// Mitsubishi GX Works2 project: 40国轩高温2次注液尝试优化   PLC: Q06UDEH (continued)
CASE iStep OF
	0:(*//初始化*)
	ConveyorMotor.xMotorCW:=0;
	ConveyorMotor.xMotorCCW:=0;
	ConveyorMotor.iProductCategoryOut:=0;
(*	//判断物料有无传感器*)	
		IF m_xPresentDelay THEN			
			ConveyorMotor.xEmpty:=0;
			IF g_xAuto AND NOT ConveyorMotor.xError THEN(*//自动情况下进行跳转*)(*无超限报警*)
				iStep:=3;
			END_IF;
		ELSE
			ConveyorMotor.xEmpty:=1;
			IF g_xAuto AND NOT ConveyorMotor.xError THEN(*//自动情况下进行跳转*)(*无超限报警*)
				iStep:=1;	
			END_IF;		
	END_IF;	
	1: (*//上料*)
	ConveyorMotor.xNextRun:=0;
	IF ConveyorMotor.xLoad    THEN (*//上料开始*)
		ConveyorMotor.iProductCategory:=0;	(*//上料开始清除产品信息*)
		iStep:=2;		
	END_IF;
	2: (*//上料完成*)
	IF ConveyorMotor.iProductCategoryIn<>0 THEN
		ConveyorMotor.iProductCategory:=ConveyorMotor.iProductCategoryIn;(* //产品信息传入*)
	END_IF;
	IF ConveyorMotor.xloadCCW THEN
		ConveyorMotor.xMotorCCW:=1; 
		ConveyorMotor.xMotorCW:=0;
	ELSE
	    ConveyorMotor.xMotorCW:=1;  
		ConveyorMotor.xMotorCCW:=0;
	END_IF;
		m_tonLoadDelay(IN:= (ConveyorMotor.xCWPresent AND NOT ConveyorMotor.xloadCCW) 
		                                        OR (ConveyorMotor.xCCWPresent AND ConveyorMotor.xloadCCW) ,
		                               PT:= ConveyorMotor.tLoadDelay ,
		                               Q:= m_xLoadDelayOut ,
		                               ET:= m_tLoadTimer );
	    IF m_xLoadDelayOut THEN 	 
		    iStep:=3;
		END_IF;
	3:(*//下料请求*)	
	ConveyorMotor.xMotorCW:=0;
	ConveyorMotor.xMotorCCW:=0;
	ConveyorMotor.xEmpty:=0;
	IF ConveyorMotor.xUnload AND NOT ConveyorMotor.xOverWidthAlarm  THEN (*无超宽报警可以下料*)
		iStep:=4;
	END_IF;
	4:(*	//下料完成*)
	IF ConveyorMotor.xUnloadCCW THEN   
		ConveyorMotor.xMotorCCW:=1;  
		ConveyorMotor.xMotorCW:=0;
		ELSE
	    ConveyorMotor.xMotorCW:=1;  
		ConveyorMotor.xMotorCCW:=0;
	END_IF;
	ConveyorMotor.xNextRun:=1; (*下一段线体旋转*)
	ConveyorMotor.iProductCategoryOut:=ConveyorMotor.iProductCategory;(*产品型号输出给下一段线体*)
	IF NOT ConveyorMotor.xUnload THEN 
		istep:=0;
	END_IF;
END_CASE;
(*In-feed zone clear and ready to accept a load from Upstream Conveyor*)
IF ldp(TRUE,g_xAuto) THEN
	m_xAutoClear:=1;
END_IF;
IF ldf(TRUE,g_xAuto) THEN
	m_xAutoClear:=0;
END_IF;
m_tonZoneClear(IN:= m_xAutoClear AND ConveyorMotor.xZoneClear ,PT:= ConveyorMotor.tZoneClearTime ,Q:=m_xZoneClearDone ,ET:= m_tZoneClearCurrentTime );
IF  m_xAutoClear AND ConveyorMotor.xZoneClear THEN
		ConveyorMotor.xMotorCW:=1; 
		iStep:=0;
END_IF;
IF ldf(TRUE, m_xAutoClear )THEN
	ConveyorMotor.xMotorCW:=0; 
END_IF;
IF NOT m_xAutoClear OR m_xZoneClearDone OR m_xPresentDelay THEN
	 m_xAutoClear:=0;
END_IF;	 
(*投入上料，搬出下料，也可用来初始化*)
IF LDP(TRUE,ConveyorMotor.xPutInto) THEN
	iStep:=0;
END_IF;
(*//当前任务显示*)
IF LDP(TRUE,ConveyorMotor.iDeviceID=g_iDeviceIDSelect) THEN
	g_iInsertTask:=ConveyorMotor.iProductCategory;
END_IF;
	(*//插入任务*)
IF g_xInsertTask AND ConveyorMotor.iDeviceID=g_iDeviceIDSelect THEN
	ConveyorMotor.iProductCategory:=g_iInsertTask;
END_IF;
(*//单线体复位，当设备号与本线体一致的时候执行复位*)
IF (g_xResetSingle AND ConveyorMotor.iDeviceID=g_iDeviceIDSelect)THEN (* //非正常情况下切断xNextRun不会复位，通过这个标志位会出发报警*)(*增加单体复位*)
	iStep:=0;
	ConveyorMotor.xNextRun:=0; 
	ConveyorMotor.xLimitAlarrm:=0;
	ConveyorMotor.xOverWidthAlarm:=0;
END_IF;
(*//手动*)
IF g_xManual THEN
(*	iStep:=0; *)(*//手动后上下料程序步骤清零*)
	(*//正转*)
	IF ConveyorMotor.xForward 
		AND ConveyorMotor.xBackward=0 
		AND ConveyorMotor.xMotorCCW=0 
		AND g_xEStop THEN
		ConveyorMotor.xMotorCW:=1;
		ConveyorMotor.xMotorCCW:=0;
		ELSE
		ConveyorMotor.xMotorCW:=0;
	END_IF;
	(*//反转*)
	IF ConveyorMotor.xBackward 
		AND ConveyorMotor.xForward=0 
		AND ConveyorMotor.xMotorCW=0 
		AND g_xEStop THEN
		ConveyorMotor.xMotorCCW:=1;
		conveyormotor.xMotorCW:=0;
		ELSE
		ConveyorMotor.xMotorCCW:=0;
	END_IF;
END_IF;
(*暂停*)
IF g_xPause THEN
	ConveyorMotor.xMotorCCW:=0;
	ConveyorMotor.xMotorCW:=0;
END_IF;
(*工作中信号输出*)
ConveyorMotor.xBusy:=ConveyorMotor.xMotorCCW OR ConveyorMotor.xMotorCW;
(*//未到达报警*)
m_tonNotArriveAlarm(IN:= iStep=0 AND ConveyorMotor.xNextRun  ,PT:= T#2s,Q:= ConveyorMotor.xNotArriveAlarm ,ET:= m_tNotArriveCurrentTime );
(*//下料超时报警*)
m_tonUnloadAlam(IN:= iStep=4,PT:=ConveyorMotor.tUnloadAlarmDelay,Q:= ConveyorMotor.xUnloadAlarm,ET:=m_tUnloadTimer );
(*//限位报警,进料检测开关失效*)
IF ( ((ConveyorMotor.xloadCCW AND NOT ConveyorMotor.xNegLimit)            (*反转上料，碰到负限位*)
	OR  ( NOT ConveyorMotor.xloadCCW AND NOT ConveyorMotor.xPosLimit)) (*正转上料，碰到正限位*)
    AND iStep=2) (*上料过程*)
    OR
   ( iStep=4 (*下料过程*)
	AND( (ConveyorMotor.xUnloadCCW AND NOT ConveyorMotor.xPosLimit)  
	OR (NOT ConveyorMotor.xUnloadCCW AND NOT ConveyorMotor.xNegLimit)))    
    THEN
    ConveyorMotor.xLimitAlarrm:=1;
    iStep:=0;
END_IF;
(*//超宽报警*)
IF (iStep=3 OR iStep=1) AND (NOT ConveyorMotor.xNegLimit OR NOT ConveyorMotor.xPosLimit) THEN
	ConveyorMotor.xOverWidthAlarm:=1;
END_IF;
(*//尺寸不足报警*)
(*//有料状态下检测两个开关都要有信号*)
IF iStep=3 AND ConveyorMotor.xSizeDeficientDetect AND (NOT ConveyorMotor.xCCWPresent OR NOT ConveyorMotor.xCWPresent)  THEN
	   ConveyorMotor.xOverWidthAlarm:=1;
	    iStep:=0;               
END_IF;
(*//总报警*)
ConveyorMotor.xError:=ConveyorMotor.xLimitAlarrm
                                              OR ConveyorMotor.xNotArriveAlarm
                                              OR ConveyorMotor.xUnloadAlarm                                             
                                              OR ConveyorMotor.xOverWidthAlarm;

(*//状态输出*)(*状态显示，容易造成指针容量不足*)
IF ConveyorMotor.xEmpty AND NOT ConveyorMotor.xBusy THEN
	m_wStateWord:=0;
END_IF;
IF ConveyorMotor.xEmpty=0 THEN
		m_wStateWord:=1;
END_IF;
IF ConveyorMotor.xBusy THEN
		m_wStateWord:=2;
END_IF;
IF ConveyorMotor.xLimitAlarrm THEN
		m_wStateWord:=3;
END_IF;
IF ConveyorMotor.xOverWidthAlarm THEN
		m_wStateWord:=4;
END_IF;
IF ConveyorMotor.xNotArriveAlarm THEN	
		m_wStateWord:=5;
END_IF;
IF ConveyorMotor.xUnloadAlarm THEN
		m_wStateWord:=6;	
END_IF;
(*选择本线体后，将状态赋值给全局变量进行显示*)
IF ConveyorMotor.iDeviceID=g_iDeviceIDSelect THEN
	g_iConveyorStatus:=m_wStateWord;
END_IF;
END_FUNCTION_BLOCK

FUNCTION_BLOCK ShuttleCar
VAR_IN_OUT
  ShuttleCarInOut : ShuttleCarIO;
END_VAR
VAR
  m_tonBrakeDelay : TON;  (* 延时 *)
  m_tBrakeDelayCurrentTime : TIME;
  m_tonArriveDelay : TON;  (* 到达延时计时器 *)
  m_xArriveDelay : BOOL;  (* 到达延时 *)
  m_tArriveDelayCurrentTime : TIME;  (* 到达延时当前时间 *)
  m_xInit : BOOL;  (* 初始化标志位 *)
  m_tonPauseDelay : TON;  (* 暂停减速 *)
  m_tPauseDelayCurrentTime : TIME;  (* 暂停延时当前时间 *)
  m_tonOvertimeAlarm : TON;  (* 超时报警定时器 *)
  m_tOvertimeCurrentTime : TIME;  (* 超时报警当前时间 *)
END_VAR
(*******************************************************************
输送小车程序，可用于使用认址片控制位置的输送车程序，可用于控制提升机，
使用了限位捕捉程序防止小车惯性过大冲过限位后继续行走，捕捉程序采用反
转复位，这样设计有弊端可能反转复位后车的位置并没有回到限位以内,当两个
限位同时碰到的时候，会使运料小车进入死锁状态，通过xPassLimit来解开死锁，
可以在触摸屏中使用一个带权限的按钮来进行控制，配合ShuttleCarCurrentPos
函数来计算位置信息
增加自动开始后将当前位置置为零的信号防止设备停在两个位置开关的中间
修改信息  修改后请增加版本
2018-1-22增加到位延时：到位延时时间可以设置，适应双向到位的位置开关，通过调整延时时间让穿梭车停在到位开关的中间
增加气缸控制信号 ShuttleCarInOut.xCylinder
增加抱闸延时 ShuttleCarInOut.tBrakeDelay
增加超时报警 ShuttleCarInOut.xOvertimeAlarm
YAO      V1.0
2018-1-22 YAO V1.1
2018-6-3：增加点动xMoveStep，单体报警复位
接口说明：
输入：
xReady    准备就绪信号，接变频器的准备就绪，无准备就绪信号的设备常置1
xForward   手动 正转
xBackward 手动 反转
iCurrentPos 当前位置信息，由外部函数给出
iDestinationPos  目标位置，自动情况下判断目标位置和当前位置的差，选择前进或后退
xPosLimit 正方向限位  常闭信号
xNegLimit 反方向限位  常闭信号
xMDIExe   自动行走使能
xPassLimit 限位屏蔽
tArriveDelay 到位延时时间设置，当前位置等于目标位置后延时相应时间后停止，默认为0
xCylinder 如果是气缸的把这个标志位置为1，
tBrakeDelay 打开抱闸延时，默认100ms。行走后会延时相应的时间打开抱闸，防止提升轴的掉落
xLooseDetect 松绳检测开关
输出：
xCW 正转输出
xCCW 反转输出
xBrake 抱闸输出 
xMDIDone 自动行走完成信号
xPosLimitCatch 正限位报警
xNegLimitCatch 负限位报警
xBusy 工作中信号
xLooseAlarm 松绳报警，报警后不可以下降，提升后如果没有松绳检测开关后复位报警信号


********************************************************************)
IF NOT m_xInit THEN
	ShuttleCarInOut.tArriveDelay:=T#0s;   (*到位延时初始化为0*)
	ShuttleCarInOut.tBrakeDelay:=T#100ms;(*抱闸延时初始化为100ms*)
	ShuttleCarInOut.tSetOverTime:=T#60s;(*超时报警初始化为1分钟*)
	m_xInit:=1;
END_IF;
(*如果是气缸的话屏蔽限位和Ready信号*)
IF ShuttleCarInOut.xCylinder THEN
	ShuttleCarInOut.xPosLimit:=1;
	ShuttleCarInOut.xNegLimit:=1;
	ShuttleCarInOut.xReady:=1;
END_IF;
(*限位捕捉，防止冲过限位开关，反转后复位*)
ShuttleCarInOut.xPosLimitCatch:=LDF(TRUE,ShuttleCarInOut.xPosLimit) OR ShuttleCarInOut.xPosLimitCatch;
IF ShuttleCarInOut.xCCW THEN  
	ShuttleCarInOut.xPosLimitCatch:=0;
END_IF;

ShuttleCarInOut.xNegLimitCatch:=LDF(TRUE,ShuttleCarInOut.xNegLimit) OR ShuttleCarInOut.xNegLimitCatch;
(*松绳报警*)
IF LDP(TRUE,ShuttleCarInOut.xLooseDetect) THEN	
	ShuttleCarInOut.xLooseAlarm:=1;
END_IF;
(*提升复位报警*)
IF ShuttleCarInOut.xCW AND NOT  ShuttleCarInOut.xLooseDetect THEN   
	ShuttleCarInOut.xLooseAlarm:=0; 
END_IF;

IF ShuttleCarInOut.xCW THEN   
	ShuttleCarInOut.xNegLimitCatch:=0; 
END_IF;

IF ShuttleCarInOut.xPassLimit OR
	g_xReset OR   (*增加复位按钮*)
	(ShuttleCarInOut.xNegLimitCatch 
	AND ShuttleCarInOut.xPosLimitCatch)  THEN  
	ShuttleCarInOut.xNegLimitCatch:=0; 
	ShuttleCarInOut.xPosLimitCatch:=0;
	ShuttleCarInOut.xLooseAlarm:=0;
END_IF;
IF ShuttleCarInOut.xReady AND g_xEStop THEN
(*手动*)
    IF g_xManual THEN  
	    IF ShuttleCarInOut.xForward 
			AND ShuttleCarInOut.xBackward=0 
			AND ShuttleCarInOut.xCCW=0 
			AND ShuttleCarInOut.xPosLimitCatch=0  THEN
		    ShuttleCarInOut.xCW:=1;
		    ELSE
		    ShuttleCarInOut.xCW:=0;
	    END_IF;
	    IF ShuttleCarInOut.xBackward 
			AND ShuttleCarInOut.xForward=0 
			AND ShuttleCarInOut.xCW=0 
			AND ShuttleCarInOut.xNegLimitCatch=0 
			AND ShuttleCarInOut.xLooseAlarm=0
			AND G_xEStop THEN  
		    ShuttleCarInOut.xCCW:=1;
		    ELSE
		    ShuttleCarInOut.xCCW:=0;
	    END_IF;
    END_IF;
    (**********)
(*自动*)
  IF g_xAuto OR ShuttleCarInOut.xMoveStep   THEN  
  	(*点动*)
  	IF LDP(TRUE,ShuttleCarInOut.xMoveStep)  THEN (*点动模式后把当前位置赋值给目标位置，防止误动作*)
  		ShuttleCarInOut.iDestinationPos:=ShuttleCarInOut.iCurrentPos;
  		END_IF;
 		IF LDP(TRUE,ShuttleCarInOut.xForward) AND ShuttleCarInOut.xMoveStep THEN
 			ShuttleCarInOut.xMDIExe:=1;
			ShuttleCarInOut.iDestinationPos:=ShuttleCarInOut.iCurrentPos+1;
		END_IF;
		IF LDP(TRUE,ShuttleCarInOut.xBackward) AND ShuttleCarInOut.xMoveStep AND ShuttleCarInOut.iCurrentPos>0  THEN
			ShuttleCarInOut.xMDIExe:=1;
			ShuttleCarInOut.iDestinationPos:=ShuttleCarInOut.iCurrentPos-1;
		END_IF;	 
	(*>>>>>>>>>>>>>>>>>>>>>>>>>>>>>>>>>>>>>*)	
	  IF ShuttleCarInOut.xMDIExe AND ShuttleCarInOut.iDestinationPos<>0 THEN	
	    IF ShuttleCarInOut.iCurrentPos<ShuttleCarInOut.iDestinationPos AND ShuttleCarInOut.xPosLimitCatch=0 THEN   (*正转*)
			ShuttleCarInOut.xCW:=1;
			ShuttleCarInOut.xCCW:=0;
			ShuttleCarInOut.xMDIDone:=0;
		END_IF;

		IF ShuttleCarInOut.iCurrentPos>ShuttleCarInOut.iDestinationPos AND ShuttleCarInOut.xNegLimitCatch=0 AND ShuttleCarInOut.xLooseAlarm=0 THEN   (*反转*)
			ShuttleCarInOut.xCCW:=1;
			ShuttleCarInOut.xCW:=0;
			ShuttleCarInOut.xMDIDone:=0;
		END_IF;
	m_tonArriveDelay(IN:= ShuttleCarInOut.iCurrentPos=ShuttleCarInOut.iDestinationPos ,
	                                    PT:= ShuttleCarInOut.tArriveDelay ,
	                                    Q:= m_xArriveDelay ,
	                                    ET:= m_tArriveDelayCurrentTime);
	     (*到位延时时间可以设置，适应双向到位的位置开关，通过调整延时时间让穿梭车停在到位开关的中间*)
		IF m_xArriveDelay AND NOT ShuttleCarInOut.xCylinder THEN
			ShuttleCarInOut.xCW:=0;
			ShuttleCarInOut.xCCW:=0;
			ShuttleCarInOut.xMDIDone:=1;
			ELSE
			ShuttleCarInOut.xMDIDone:=0;
		END_IF;

		IF ShuttleCarInOut.xPosLimitCatch THEN
			ShuttleCarInOut.xCW:=0;
			ShuttleCarInOut.xMDIDone:=0;
		END_IF;

		IF ShuttleCarInOut.xNegLimitCatch  OR ShuttleCarInOut.xLooseAlarm THEN
			ShuttleCarInOut.xCCW:=0;
			ShuttleCarInOut.xMDIDone:=0;
		END_IF;
		ELSE(*MDIExe AND DestinationPos<>0的ELSE*)
		ShuttleCarInOut.xCW:=0;
		ShuttleCarInOut.xCCW:=0;
		ShuttleCarInOut.xMDIDone:=0;
	  END_IF;
	END_IF;
	ELSE  (*无就绪信号   或急停的情况下*)
		ShuttleCarInOut.xCW:=0;
		ShuttleCarInOut.xCCW:=0;	
END_IF;
    (*抱闸延时*)
m_tonBrakeDelay(IN:= ShuttleCarInOut.xCW OR ShuttleCarInOut.xCCW,
                                    PT:= ShuttleCarInOut.tBrakeDelay,
                                    Q:=ShuttleCarInOut.xBrake ,
                                    ET:= m_tBrakeDelayCurrentTime);

(*自动上电后把当前位置清零，防止穿梭车不在开关位置*)
(**------这里增加MDIexe上升沿是因为有时目标地址是2，但MDI没有了就会往下掉，导致当前位置还是2，却不在开关位置，无法上下料**)
(*程序这么写就意味着必须上为2，下为1*)
IF LDP(TRUE,g_xAuto ) OR NOT ShuttleCarInOut.xMDIExe THEN
	ShuttleCarInOut.iCurrentPos:=0;
END_IF;
IF ShuttleCarInOut.xCW OR ShuttleCarInOut.xCCW THEN
	ShuttleCarInOut.xBusy:=1;
	ELSE
	ShuttleCarInout.xBusy:=0;
END_IF;

(*暂停，带延时减速斜坡，ShuttleCarInOut.xPauseRamp为减速斜坡输出位*)
m_tonPauseDelay(IN:=g_xPause,PT:= T#2s ,Q:=ShuttleCarInOut.xPauseRamp,ET:= m_tPauseDelayCurrentTime );
IF ShuttleCarInOut.xPauseRamp THEN
	ShuttleCarInOut.xCW:=0;
	ShuttleCarInOut.xCCW:=0;
	ShuttleCarInOut.xBrake:=0;
END_IF;
(*超时报警*)
m_tonOvertimeAlarm(IN:= ShuttleCarInOut.xMDIExe AND (ShuttleCarInOut.iCurrentPos<>ShuttleCarInOut.iDestinationPos) ,
                                           PT:= ShuttleCarInOut.tSetOverTime,
                                           Q:= ShuttleCarInOut.xOvertimeAlarm ,
                                           ET:= m_tOvertimeCurrentTime );
(*//单体复位，当设备号与本设备一致的时候执行复位*)
IF (g_xResetSingle AND ShuttleCarInOut.diDeviceID=g_diDeviceIDSelect)THEN(*增加单体复位*)
	ShuttleCarInOut.iCurrentPos:=0;
END_IF;
END_FUNCTION_BLOCK

FUNCTION_BLOCK Switch
VAR_IN_OUT
  ConveyorEntryIO : ConveyorIO;
  ConveyorExitIO : ConveyorIO;
END_VAR
VAR
  m_tonLiftCylinderDelay : TON;  (* 顶升延时 *)
  m_xLiftCylinderDelay : BOOL;
  m_tLiftCylinderDelay : TIME;
  m_tonExitBarDelay : TON;  (* 退出阻挡器延时 *)
  m_tExitBarDelay : TIME;
  m_xExitBarDelay : BOOL;
END_VAR
VAR_IN_OUT
  SwitchIO : SwitchIO;
END_VAR
VAR
  iStep : INT;
  m_xInitial : BOOL;
  m_tonCylinderOvertime : TON;  (* 气缸超时报警定时器 *)
  m_tCylinderOvertimeCurrent : TIME;
END_VAR
(**************************************************
//顶升移载模块，抽象为一条输入输线 ，一条输出输送线
//一个进入阻挡器，一个放出阻挡器，和一个顶升气缸的控制
//程序思路比较混乱，接口不清晰，需要整改
//直接放行的时候有问题
//switchEnable =0的时候   离开线体的PutInto有问题
//增加xPutInto程序
//12-17日   V1.0
//***************************************************)
(*ConveyorEntry(ConveyorMotor:=ConveyorEntryIO);
(*ConveyorExit(ConveyorMotor:=ConveyorExitIO);*)


IF NOT m_xInitial THEN
	SwitchIO.tSetOvertime:=T#5s;
	SwitchIO.xExitEnable:=1;
	m_xInitial:=1;
END_IF;
IF g_xAuto THEN
	CASE iStep OF
		0:(*初始化*)
		ConveyorEntryIO.xLoad:=0;
		ConveyorEntryIO.xUnload:=0;
		ConveyorEntryIO.xPutInto:=0;
		ConveyorExitIO.xLoad:=0;
		ConveyorExitIo.xUnload:=0;
		ConveyorExitIO.xPutInto:=0;
		SwitchIO.xEntryBarCylinderRetract:=0;
		SwitchIO.xExitBarCylinderRetract:=0;
		IF SwitchIO.xLiftCylinderExtendInit THEN
			SwitchIO.xLiftCylinderExtend:=1;
			SwitchIO.xLiftCylinderRetract:=0;
		    IF SwitchIO.xLiftCylinderExtendDetect THEN
			    iStep:=1;
			END_IF; 
			ELSE
			SwitchIO.xLiftCylinderExtend:=0;
			SwitchIO.xLiftCylinderRetract:=1;	
		    IF SwitchIO.xLiftCylinderRetractDetect THEN
			    iStep:=1;
		    END_IF;		
		END_IF;
		1:(*上料*)
        IF SwitchIO.xEntryEnable AND ConveyorEntryIO.xEmpty AND ConveyorExitIO.xEmpty THEN
        	SwitchIO.xEntryBarCylinderRetract:=1;
        	ConveyorEntryIO.xLoad:=1;
        END_IF;
        IF ConveyorEntryIO.xEmpty=0 THEN
        	SwitchIO.xEntryBarCylinderRetract:=0;
        	ConveyorEntryIO.xLoad:=0;
        	ConveyorExitIO.xPutInto:=ConveyorExitIO.xEmpty;
        END_IF;
        SwitchIO.xExitBarCylinderRetract:=NOT SwitchIO.xSwithEnable;
        IF m_xLiftCylinderDelay AND  SwitchIO.xSwithEnable AND SwitchIO.xExitEnable THEN
			iStep:=2;
        END_IF;
        IF SwitchIO.xSwithEnable=0 AND m_xLiftCylinderDelay AND SwitchIO.xExitEnable  THEN
			iStep:=3;
        END_IF;
		2:(*顶升*)
		ConveyorExitIO.iProductCategory:=ConveyorEntryIO.iProductCategory;
		ConveyorExitIO.iTaskID:=ConveyorEntryIO.iTaskID;
		ConveyorExitIO.diDesConveyor:=ConveyorEntryIO.diDesConveyor;
		SwitchIO.xExitBarCylinderRetract:=0;
		ConveyorExitIO.xPutInto:=0;
		IF SwitchIO.xLiftCylinderExtendInit THEN
			SwitchIO.xLiftCylinderExtend:=0;
			SwitchIO.xLiftCylinderRetract:=1;
		    ELSE
			SwitchIO.xLiftCylinderExtend:=1;
			SwitchIO.xLiftCylinderRetract:=0;			
		END_IF;

		IF SwitchIO.xLiftCylinderExtendInit THEN
		  	IF SwitchIO.xLiftCylinderRetractDetect THEN
		  		iStep:=4;
		  	END_IF;
		  	ELSE
		  	IF SwitchIO.xLiftCylinderExtendDetect THEN
				iStep:=4; 
		  	END_IF;
		END_IF;
		3:(*放行*)	
		ConveyorExitIO.iProductCategory:=ConveyorEntryIO.iProductCategory;
		ConveyorExitIO.iTaskID:=ConveyorEntryIO.iTaskID;
		ConveyorExitIO.diDesConveyor:=ConveyorEntryIO.diDesConveyor;
		ConveyorExitIO.xPutInto:=0;
		iStep:=4;
		4:(*下料*)
		(*通过出料传输线下料*)
		IF SwitchIO.xExitEnable  AND m_xExitBarDelay AND NOT SwitchIO.xExitBarCylinderRetract  THEN		  
		  	ConveyorExitIO.xUnload:=1;
			ELSE
		  	ConveyorExitIO.xUnload:=0;
		END_IF;	
		(*通过进料传输线下料*)
		IF SwitchIO.xExitEnable  AND m_xExitBarDelay  AND SwitchIO.xExitBarCylinderRetract THEN		  
		  	ConveyorEntryIO.xUnload:=1;
			ELSE
		  	ConveyorEntryIO.xUnload:=0;
		END_IF;			    	
		IF (ConveyorExitIO.xEmpty OR ConveyorEntryIO.xEmpty) AND m_xExitBarDelay  THEN
		  	ConveyorExitIO.xPutInto:=1;
		  	ConveyorEntryIO.xPutInto:=1;
			iStep:=0; 
		END_IF;
	END_CASE;
	m_tonLiftCylinderDelay(IN:=NOT ConveyorEntryIO.xEmpty AND iStep=1 ,PT:= T#1S ,Q:= m_xLiftCylinderDelay ,ET:=m_tLiftCylinderDelay );
	m_tonExitBarDelay(IN:=iStep=4 ,PT:= T#1s ,Q:= m_xExitBarDelay ,ET:= m_tExitBarDelay);
END_IF;
(*复位程序*)
IF (g_xResetSingle AND  (g_diDeviceIDSelect=ConveyorEntryIO.diDeviceID OR g_diDeviceIDSelect=ConveyorExitIO.diDeviceID))
	OR LDP(TRUE,SwitchIO.xLiftCylinderExtendInit) 
	OR LDF(TRUE,SwitchIO.xLiftCylinderExtendInit) 
	OR LDP(TRUE,SwitchIO.xPutInto)  THEN
	ConveyorEntryIO.xPutInto:=1;
	ConveyorExitIO.xPutInto:=1;
	iStep:=0;
END_IF;

IF g_xManual  THEN
	iStep:=0;
	ConveyorEntryIO.xLoad:=0;
    ConveyorEntryIO.xUnload:=0;
	ConveyorEntryIO.xPutInto:=0;
	ConveyorExitIO.xLoad:=0;
	ConveyorExitIo.xUnload:=0;
	ConveyorExitIO.xPutInto:=0;
	SwitchIO.xEntryBarCylinderRetract:=0;
	SwitchIO.xExitBarCylinderRetract:=0;
	IF SwitchIO.xEntryBarCylinderRetractButton THEN
		SwitchIO.xEntryBarCylinderRetract:=1;
		ELSE
		SwitchIO.xEntryBarCylinderRetract:=0;
	END_IF;
	IF SwitchIO.xExitBarCylinderRetractButton THEN
		SwitchIO.xExitBarCylinderRetract:=1;
		ELSE
		SwitchIO.xExitBarCylinderRetract:=0;
	END_IF;
	IF SwitchIO.xLiftCylinderExtendButton AND NOT SwitchIO.xLiftCylinderRetractButton THEN
		SwitchIO.xLiftCylinderExtend:=1;
		SwitchIO.xLiftCylinderRetract:=0;
	END_IF;
	IF NOT SwitchIO.xLiftCylinderExtendButton AND  SwitchIO.xLiftCylinderRetractButton THEN
		SwitchIO.xLiftCylinderExtend:=0;
		SwitchIO.xLiftCylinderRetract:=1;
	END_IF;		 
END_IF;
(*气缸超时报警*)
m_tonCylinderOvertime(IN:= (SwitchIO.xLiftCylinderExtend AND NOT SwitchIO.xLiftCylinderExtendDetect) 
OR  (SwitchIO.xLiftCylinderRetract AND NOT SwitchIO.xLiftCylinderRetractDetect) ,
PT:= SwitchIO.tSetOvertime ,Q:= SwitchIO.xOvertimeAlarm ,ET:= m_tCylinderOvertimeCurrent );
END_FUNCTION_BLOCK

FUNCTION_BLOCK PreemptivePriority
VAR_INPUT
  xCondition : ARRAY [1..13] OF BOOL;  (* 条件1 *)
  xTaskComplete : BOOL;  (* 任务完成 *)
  xReset : BOOL;  (* 复位 *)
END_VAR
VAR
  xOccupy : BOOL;  (* 占用 *)
END_VAR
VAR_OUTPUT
  iPriority : INT;  (* 输出任务号 *)
END_VAR
VAR
  m_tonConditionDelay : TON;
  m_xConditionDelay : BOOL;
  m_tConditionCurrentTime : TIME;
  m_iLastTask : INT;  (* 上次执行的任务 *)
  m_tpLastTaskPulse1 : TP;
  m_tpLastTaskPulse2 : TP;
  m_tpLastTaskPulse3 : TP;
  m_tpLastTaskPulse4 : TP;
  m_tpLastTaskPulse5 : TP;
  m_xLastTaskPulse : ARRAY [1..13] OF BOOL;
  m_tLastTaskPulse : ARRAY [1..13] OF TIME := [13(T#0s)];
  m_tpLastTaskPulse6 : TON;
  ii : INT;
END_VAR
VAR CONSTANT
  CONDITION_QUANTITY : INT := 13;
END_VAR
VAR
  m_tpLastTaskPulse7 : TON;
  m_tpLastTaskPulse8 : TON;
  m_tpLastTaskPulse9 : TON;
  m_tpLastTaskPulse10 : TON;
  m_tpLastTaskPulse11 : TON;
  m_tpLastTaskPulse12 : TON;
  m_tpLastTaskPulse13 : TON;
END_VAR
(*抢占式优先级块
现在满足13个条件的任务进行抢占式优先级排列
条件满足后延时两秒，开始执行任务，
同一任务连续执行优先级下降
需要改造成任意多个
使用于一个入口多个出口的程序，使用抢占式优先级块
*)
IF LDP(TRUE, xTaskComplete) THEN
	xOccupy:=0;
	iPriority:=0;
END_IF;
(*//任务滤波，延时两秒*)
m_tonConditionDelay(IN:=( xCondition[1]
						OR xCondition[2]
						OR xCondition[3]
						OR xCondition[4]
						OR xCondition[5]
						OR xCondition[6]
						OR xCondition[7]
						OR xCondition[8]
						OR xCondition[9]
						OR xCondition[10]
						OR xCondition[11]
						OR xCondition[12]
						OR xCondition[13]
						)
						AND iPriority=0,
					PT:= T#1s,
					Q:= m_xConditionDelay ,
					ET:= m_tConditionCurrentTime );		
(*//判断优先级，上个任务与本次任务相同，延时一秒执行*)
m_tpLastTaskPulse1(IN:= xCondition[1]  AND m_iLastTask=1 AND m_xConditionDelay  ,PT:= T#1s,Q:= m_xLastTaskPulse[1],ET:= m_tLastTaskPulse[1] );
m_tpLastTaskPulse2(IN:= xCondition[2]  AND m_iLastTask=2 AND m_xConditionDelay  ,PT:= T#1s,Q:= m_xLastTaskPulse[2],ET:= m_tLastTaskPulse[2] );
m_tpLastTaskPulse3(IN:= xCondition[3]  AND m_iLastTask=3 AND m_xConditionDelay  ,PT:= T#1s,Q:= m_xLastTaskPulse[3],ET:= m_tLastTaskPulse[3] );
m_tpLastTaskPulse4(IN:= xCondition[4]  AND m_iLastTask=4 AND m_xConditionDelay  ,PT:= T#1s,Q:= m_xLastTaskPulse[4],ET:= m_tLastTaskPulse[4] );
m_tpLastTaskPulse5(IN:= xCondition[5]  AND m_iLastTask=5 AND m_xConditionDelay  ,PT:= T#1s,Q:= m_xLastTaskPulse[5],ET:= m_tLastTaskPulse[5] );
m_tpLastTaskPulse6(IN:= xCondition[6]  AND m_iLastTask=6 AND m_xConditionDelay  ,PT:= T#1s,Q:= m_xLastTaskPulse[6],ET:= m_tLastTaskPulse[6] );
m_tpLastTaskPulse7(IN:= xCondition[7]  AND m_iLastTask=7 AND m_xConditionDelay  ,PT:= T#1s,Q:= m_xLastTaskPulse[7],ET:= m_tLastTaskPulse[7] );
m_tpLastTaskPulse8(IN:= xCondition[8]  AND m_iLastTask=8 AND m_xConditionDelay  ,PT:= T#1s,Q:= m_xLastTaskPulse[8],ET:= m_tLastTaskPulse[8] );
m_tpLastTaskPulse9(IN:= xCondition[9]  AND m_iLastTask=9 AND m_xConditionDelay  ,PT:= T#1s,Q:= m_xLastTaskPulse[9],ET:= m_tLastTaskPulse[9] );
m_tpLastTaskPulse10(IN:= xCondition[10]  AND m_iLastTask=10 AND m_xConditionDelay  ,PT:= T#1s,Q:= m_xLastTaskPulse[10],ET:= m_tLastTaskPulse[10] );
m_tpLastTaskPulse11(IN:= xCondition[11]  AND m_iLastTask=11 AND m_xConditionDelay  ,PT:= T#1s,Q:= m_xLastTaskPulse[11],ET:= m_tLastTaskPulse[11] );
m_tpLastTaskPulse12(IN:= xCondition[12]  AND m_iLastTask=12 AND m_xConditionDelay  ,PT:= T#1s,Q:= m_xLastTaskPulse[12],ET:= m_tLastTaskPulse[12] );
m_tpLastTaskPulse13(IN:= xCondition[13]  AND m_iLastTask=13 AND m_xConditionDelay  ,PT:= T#1s,Q:= m_xLastTaskPulse[13],ET:= m_tLastTaskPulse[13] );
(*//执行*)
FOR ii:=1 TO CONDITION_QUANTITY BY 1 DO 
	IF NOT xCondition[ii] AND NOT xOccupy THEN
		iPriority:=0;
	END_IF;
	IF xCondition[ii] AND NOT xOccupy AND m_xConditionDelay AND NOT  m_xLastTaskPulse[ii]  THEN
		iPriority:=ii;
		xOccupy:=1;
		m_iLastTask:=ii;
	END_IF;
END_FOR;        
(*//复位*)
IF xReset THEN
	iPriority:=0;
	xOccupy:=0;
	m_iLastTask:=0;	
END_IF;
(*//清除占用*)
IF iPriority=0 THEN
	xOccupy:=0;
END_IF;
END_FUNCTION_BLOCK

FUNCTION_BLOCK PriorityQueue
VAR_INPUT
  arrxCondition : ARRAY [1..13] OF QueueElement;
  xTaskComplete : BOOL;  (* 任务完成 *)
  xReset : BOOL;  (* 复位 *)
END_VAR
VAR
  xOccupy : BOOL;  (* 占用 *)
END_VAR
VAR_OUTPUT
  iPriority : INT;  (* 输出任务号 *)
END_VAR
VAR
  jj : INT;
END_VAR
VAR CONSTANT
  CONDITION_QUANTITY : INT := 13;
END_VAR
VAR
  arriTaskStack : ARRAY [0..13] OF INT;
  ii : INT;
  kk : INT;
  arrxConditionDelay : ARRAY [1..13] OF BOOL;
  arrxConditionEdgeDetect : ARRAY [1..13] OF BOOL;
  arrxDelayEdgeDetect : ARRAY [1..13] OF BOOL;
  arriDelayCounter : ARRAY [1..13] OF INT;
  ll : INT;
  Temp : INT;
  mm : INT;
  nn : INT;
  Temp2 : INT;
  oo : INT;
END_VAR
(****************************************************************************)
(*
一般情况多对一的任务调度采用这个结构，排队通过出口
优先级功能块，存储任意条件的优先级，实现栈功能先入先出，
复位功能还有问题，
出入栈式优先级块，满足条件后入栈，先入先出，在栈尾加载新任务
栈首为当前执行的任务，任务完成使用上升沿触发，触发后栈首元素弹出

复位功能清空堆栈，栈的容量在CONDITION_QUANTITY 设置
增加了结构体，结构体中带有一个条件函数，和一个优先级指示
任务完成后通过凭借优先级来排序，优先级高的条件先执行   优先级排序是从小到大的，数值小的优先级高
防止干扰，增加了任务的1秒的延时
*)

(***************************************************************************)
(*(//入栈*)
FOR ii:=1 TO CONDITION_QUANTITY BY 1 DO
	(*//循环内无法用定时器，改用计数器的形式*)
	IF arrxCondition[ii].xCondition AND SM411 (*//0.2秒的方波信号，如果移植需要修改成两个定时器*)
		AND arriDelayCounter[ii]<6  (* //计数为6，5个0.2秒的方波，所以为1秒*)
		AND NOT arrxDelayEdgeDetect[ii] THEN    (*//循环内无法用沿函数，增加锁定标志位*)
		arriDelayCounter[ii]:=arriDelayCounter[ii]+1;   (*//计数*)
	END_IF;
	IF NOT arrxCondition[ii].xCondition THEN
		arriDelayCounter[ii]:=0;   (*//计数清零*)
	END_IF;
	arrxDelayEdgeDetect[ii]:=arrxCondition[ii].xCondition AND SM411;  (*//沿函数锁*)
	IF arriDelayCounter[ii]=5 AND NOT arrxConditionEdgeDetect[ii] THEN;  (*//条件满足1秒后*)
		FOR kk:=0 TO CONDITION_QUANTITY BY 1 DO    
			IF arriTaskStack[kk]=0 THEN
				arriTaskStack[kk]:=ii;   (*//栈尾添加*)
				EXIT;
			END_IF;		
		END_FOR;
	END_IF;	
	arrxConditionEdgeDetect[ii]:=arriDelayCounter[ii]=5;  (*//边沿*)
END_FOR;
(*//栈顶任务为当前执行的任务**)
iPriority:=arriTaskStack[0]; 
(*//栈顶任务完成，弹出*)
IF 	LDP(TRUE, xTaskComplete) THEN
	FOR jj:=0 TO CONDITION_QUANTITY-1 BY 1 DO
		arriTaskStack[jj]:=arriTaskStack[jj+1];
	END_FOR;
	arriTaskStack[CONDITION_QUANTITY]:=0;(*//栈尾清零*)
	(*//排序，使用插入排序*)
	FOR oo:=0 TO CONDITION_QUANTITY BY 1 DO
		IF arriTaskStack[oo]=0 THEN
			EXIT;  (* //寻找栈中不为零的元素  ，防止0元素进入条件查找的时候报错*)
		END_IF;
	END_FOR;
	(*//插入排序insertionsort*)
	FOR mm:=1 TO oo-1  BY 1 DO   (*//从1开始*)
		Temp:=arriTaskStack[mm];  (*//当前数据记录 *)
		Temp2:=arrxCondition[arriTaskStack[mm]].iPriority;  (*//当前优先级记录 *)
		nn:=mm;  (*//指针赋值*)
		WHILE  (nn>0 AND Temp2< arrxCondition[arriTaskStack[nn-1]].iPriority)  DO  (*//优先级比较，当前优先级小于他前面元素优先级的时候*)
			 arriTaskStack[nn] := arriTaskStack[nn-1] ;  (*//优先级低的向后复制，比TEMP2大的元素都要复制到下一个位置*)
			 nn:=nn-1;
		END_WHILE;
		arriTaskStack[nn]:=Temp; (*//把当前数据放在合适的位置*)
	END_FOR;
END_IF;
(*//复位*)
IF xReset THEN
	FOR jj:=0 TO CONDITION_QUANTITY BY 1 DO
		arriTaskStack[jj]:=0;
	END_FOR;
	FOR ll:=1 TO CONDITION_QUANTITY BY 1 DO
		arrxConditionEdgeDetect[ll]:=0;
		arriDelayCounter[ll]:=0;
	END_FOR;
END_IF;
END_FUNCTION_BLOCK

FUNCTION_BLOCK Conveyor
VAR
  m_xPresentDelay : BOOL;  (* 有无判断延时 *)
  m_xLoadDelayOut : BOOL;  (* 上料延时输出 *)
  m_xInitial : BOOL;  (* 初始化 *)
  m_tUnloadTimer : TIME;  (* 下料计时器 *)
  m_tPresentDelayCurrentTime : TIME;
  m_tonUnloadAlam : TON;  (* 下料报警定时器 *)
  m_tonPresentDelay : TON;  (* 物料有无判断延时，防止误动作 *)
  m_tonNotArriveAlarm : TON;  (* 未到达报警计时 *)
  m_tonLoadDelay : TON;  (* 上料延时 *)
  m_tNotArriveCurrentTime : TIME;  (* 未到达报警计时当前时间 *)
  m_tLoadTimer : TIME;  (* 上料计时器 *)
  iStep : INT;  (* 上料步骤 *)
  m_wStateWord : INT;
END_VAR
VAR_IN_OUT
  ConveyorMotor : ConveyorIO;  (* 输送线输入输出 *)
END_VAR
VAR
  m_tonZoneClear : TON;  (* 初始化清除 *)
  m_tZoneClearCurrentTime : TIME;  (* 初始化清除当前时间 *)
  m_xAutoClear : BOOL;  (* 初始化清除标志位 *)
  m_xZoneClearDone : BOOL;  (* 初始化清除完成 *)
END_VAR
(*////////////////////////////////////////////////////////////////////////////////////////////////////////////
//传输线控制FB块，可控制单方向线体，双向旋转线体，支持双向上下料            
//线体初始化后为空的情况下输入xLoad信号即可进行上料动作，使用xLoadCCW信号可反方向上料
//增加了产品信息和产品种类的储存，当传输线为空和上料进行标志位为零的情况下清除产品信息和产品种类
//使用方式是在置位xLoad信号后，把产品信息和产品种类传入，等下料后自动清零
//线体不为空的情况下使用xUnload信号可进行下料动作，物料有无传感器的下降沿后出发计时器，延时断开传输线旋转
//单方向传输线体把xLoadCCW、xUnloadCCW设置为零，双向线体上料方向和下料反向的,方向固定的 把xUnloadCCW设置为1
//双方向线体双向都能上下料的要根据上料的方向来设置xLoadCCW,xUnloadCCW
//增加工作中信号xBusy当电机正转 显示为工作中
//增加上下料超时报警，xLoadAlarm，xUnloadAlarm，设定时间在LOAD_UNLOAD_TIME常量上，现在设置的为30秒
//增加xPutInto信号，用于直接投入的物料，检测开关感应到后，直接进入下料流程，上升沿有效
//离开延时改为变量 iLeaveDelay 默认为0 离开检测开关离输送线尾端比较远的线体需要根据情况设定100ms为单位
//增加初始化标志位，增加进入延时时间，初始化为进入延时时间为0 ，离开延时时间为2S，通过外围接口可以更改
//修改信息  修改后请增加版本
//12-17进行了优化，增加了未到达报警，当物料未传送到下一设备，就报未到达报警，使用xNextRun标志位制作，没有正常到达
//第0步，不能跳转到第一步把标志位复位，即出现中断情况，2秒后报警
//修改信息  修改后请增加版本
//上料延时增加为50ms防止干扰信号
//nextrun信号在 第三步也要复位
//增加限位报警
//增加超宽报警
//增加产品型号输出在下料的时候把产品型号输送给下一段线体
//增加线体单独复位
//增加任务插入功能配合全局变量
//增加暂停功能
//增加线体状态字显示  0 空闲 1：有料  2 工作中  3  超限报警 4 超宽报警  5 未到达报警  6 下料超时报警
//空料判断放在自动前，进行有无报警判断，然后跳转
//修改超限报警，与尺寸检测报警
////YAO      V1.0
//把所有的IF语句去掉，  IF语句占用指针存储区，容易造成存储区不足的现象
////YAO      V1.1
//初始化清除线体标志位xZoneClear
//ZPA zero pressure accumulation  Term that describes the Conveyor controls and mechanical scheme that will 
//cause loads to queue on a conveyor in discrete zones such that loads do not touch each other(wrapped boxed tray tote carton)
//除了产品信息外，还增加了目标地址，任务类型的数据传递。
//YAO      V1.0
///////////////////////////////////////////////////////////////////////////////////////////////////////////
(*********************************************************)
(*//初始化，
//上料延时位0S，下料报警延时为30S
//下料延时设一个比较大的时间，主要依靠xunload标志位来停止输送线，特殊情况可以用延时来停止物流线下料
//设置时间大的时候计时器会失效*)
IF NOT m_xInitial THEN
	ConveyorMotor.tLoadDelay:=T#100ms;
	ConveyorMotor.tUnloadAlarmDelay:=T#30s;
	ConveyorMotor.xPosLimit:=1;
	ConveyorMotor.xNegLimit:=1;
	ConveyorMotor.xSizeDeficientDetect:=0;
	ConveyorMotor.xZoneClear:=0;
	ConveyorMotor.tZoneClearTime:=T#10s;
	m_xInitial:=1;
END_IF;
(*//自动
//复位信号把步号置0，但xLoad与xUnload没有复位，调用程序需要注意复位后把这两个信号置零，以免发生误动作
//物料有无判断增加延时，防止开自动瞬间误动作发生*)
m_tonPresentDelay(IN:= ConveyorMotor.xCWPresent OR ConveyorMotor.xCCWPresent,
					PT:=T#100ms,
					Q:= m_xPresentDelay,
					ET:= m_tPresentDelayCurrentTime);
CASE iStep OF
0:(*//初始化*)
	ConveyorMotor.xMotorCW:=0;
	ConveyorMotor.xMotorCCW:=0;
	ConveyorMotor.xNextRun:=0;
	ConveyorMotor.iProductCategoryOut:=0;
	ConveyorMotor.iTaskIDOut:=0;
	ConveyorMotor.diDesConveyorOut:=0;
	out(NOT m_xPresentDelay,ConveyorMotor.xEmpty);(*	//判断物料有无传感器*)	
	mov(m_xPresentDelay AND g_xAuto AND NOT ConveyorMotor.xError,3,iStep);(*//自动情况下进行跳转*)(*无超限报警*)
	mov(NOT m_xPresentDelay AND g_xAuto AND NOT ConveyorMotor.xError,1,iStep);
1: (*//上料*)
	rst(ConveyorMotor.xLoad ,ConveyorMotor.iProductCategory);(*//上料开始清除产品信息*)
	rst(ConveyorMotor.xLoad ,ConveyorMotor.iTaskID);
	rst(ConveyorMotor.xLoad ,ConveyorMotor.diDesConveyor);
	mov(ConveyorMotor.xLoad,2,iStep);
2: (*//上料完成*)
	ConveyorMotor.iProductCategory:=ConveyorMotor.iProductCategoryIn;(* //产品信息传入*)
	ConveyorMotor.iTaskID:=ConveyorMotor.iTaskIDIn;
	ConveyorMotor.diDesConveyor:=ConveyorMotor.diDesConveyorIn;
	set(ConveyorMotor.xloadCCW,ConveyorMotor.xMotorCCW);
	rst(ConveyorMotor.xloadCCW,ConveyorMotor.xMotorCW);
	set(NOT ConveyorMotor.xloadCCW,ConveyorMotor.xMotorCW);
	rst(NOT ConveyorMotor.xloadCCW,ConveyorMotor.xMotorCCW);	
	m_tonLoadDelay(IN:= (ConveyorMotor.xCWPresent AND NOT ConveyorMotor.xloadCCW) 
												OR (ConveyorMotor.xCCWPresent AND ConveyorMotor.xloadCCW) ,
										PT:= ConveyorMotor.tLoadDelay ,
										Q:= m_xLoadDelayOut ,
										ET:= m_tLoadTimer );
	mov(m_xLoadDelayOut,3, iStep);
3:(*//下料请求*)	
	ConveyorMotor.xMotorCW:=0;
	ConveyorMotor.xMotorCCW:=0;
	ConveyorMotor.xEmpty:=0;
	mov(ConveyorMotor.xUnload AND NOT ConveyorMotor.xOverWidthAlarm,4,iStep);
4:(*	//下料完成*)
	set(ConveyorMotor.xUnloadCCW,ConveyorMotor.xMotorCCW);
	rst(ConveyorMotor.xUnloadCCW,ConveyorMotor.xMotorCW);
	set(NOT ConveyorMotor.xUnloadCCW,ConveyorMotor.xMotorCW);
	rst(NOT ConveyorMotor.xUnloadCCW,ConveyorMotor.xMotorCCW);	
	ConveyorMotor.xNextRun:=1; (*下一段线体旋转*)
	ConveyorMotor.iProductCategoryOut:=ConveyorMotor.iProductCategory;(*产品型号输出给下一段线体*)
	ConveyorMotor.iTaskIDOut:=ConveyorMotor.iTaskID;
	ConveyorMotor.diDesConveyorOut:=ConveyorMotor.diDesConveyor;
	mov( NOT ConveyorMotor.xUnload , 0, istep );
END_CASE;
(*In-feed zone clear and ready to accept a load from Upstream Conveyor*)
set(ldp(TRUE,g_xAuto) ,m_xAutoClear);
rst(ldf(TRUE,g_xAuto) ,m_xAutoClear);
m_tonZoneClear(IN:= m_xAutoClear AND ConveyorMotor.xZoneClear ,PT:= ConveyorMotor.tZoneClearTime ,Q:=m_xZoneClearDone ,ET:= m_tZoneClearCurrentTime );
set(m_xAutoClear AND ConveyorMotor.xZoneClear,ConveyorMotor.xMotorCW);
mov( m_xAutoClear AND ConveyorMotor.xZoneClear, 0 ,iStep );
rst(  ldf(TRUE, m_xAutoClear ) ,ConveyorMotor.xMotorCW);
rst( m_xZoneClearDone OR m_xPresentDelay  , m_xAutoClear );
(*投入上料，搬出下料，也可用来初始化*)
movp( ConveyorMotor.xPutInto, 0 , iStep );
(*//当前任务显示*)
movp( ConveyorMotor.diDeviceID=g_diDeviceIDSelect , ConveyorMotor.iProductCategory , g_iInsertCategory );
movp( ConveyorMotor.diDeviceID=g_diDeviceIDSelect , ConveyorMotor.iTaskID , g_iInsertTaskID );
dmovp( ConveyorMotor.diDeviceID=g_diDeviceIDSelect , ConveyorMotor.diDesConveyor , g_diInsertDesConveyor );
(*//插入任务*)
mov(g_xInsertTask AND ConveyorMotor.diDeviceID=g_diDeviceIDSelect ,g_iInsertCategory , ConveyorMotor.iProductCategory );
mov(g_xInsertTask AND ConveyorMotor.diDeviceID=g_diDeviceIDSelect , g_iInsertTaskID , ConveyorMotor.iTaskID );
dmov(g_xInsertTask AND ConveyorMotor.diDeviceID=g_diDeviceIDSelect , g_diInsertDesConveyor , ConveyorMotor.diDesConveyor );
(*//单线体复位，当设备号与本线体一致的时候执行复位*)
mov(g_xResetSingle AND ConveyorMotor.diDeviceID=g_diDeviceIDSelect , 0 , iStep );
rst(g_xResetSingle AND ConveyorMotor.diDeviceID=g_diDeviceIDSelect ,ConveyorMotor.xNextRun );
rst(g_xResetSingle AND ConveyorMotor.diDeviceID=g_diDeviceIDSelect  ,ConveyorMotor.xLimitAlarrm );
rst(g_xResetSingle AND ConveyorMotor.diDeviceID=g_diDeviceIDSelect  ,ConveyorMotor.xOverWidthAlarm );
(*//手动*)
(*//正转*)
set( g_xManual 
AND ConveyorMotor.xForward 
AND ConveyorMotor.xBackward=0 
AND ConveyorMotor.xMotorCCW=0 
AND g_xEStop  , 
ConveyorMotor.xMotorCW);
rst((g_xManual 
AND (NOT ConveyorMotor.xForward  
OR ConveyorMotor.xBackward 
OR ConveyorMotor.xMotorCCW )) 
OR NOT g_xEStop,
ConveyorMotor.xMotorCW);
(*//反转*)		
set(g_xManual 
AND ConveyorMotor.xBackward 
AND ConveyorMotor.xForward=0 
AND ConveyorMotor.xMotorCW=0 
AND g_xEStop ,
ConveyorMotor.xMotorCCW);
rst((g_xManual AND 
(NOT ConveyorMotor.xBackward  
OR ConveyorMotor.xForward 
OR ConveyorMotor.xMotorCW ) ) 
OR NOT g_xEStop,
ConveyorMotor.xMotorCCW);
mov(g_xManual ,0,iStep);(*//手动后上下料程序步骤清零*)
(*暂停*)
rst(g_xPause,ConveyorMotor.xMotorCCW);
rst( g_xPause , ConveyorMotor.xMotorCW );
(*工作中信号输出*)
ConveyorMotor.xBusy:=ConveyorMotor.xMotorCCW OR ConveyorMotor.xMotorCW;
(*//未到达报警*)
m_tonNotArriveAlarm(IN:= iStep=0 AND ConveyorMotor.xNextRun  ,PT:= T#2s,Q:= ConveyorMotor.xNotArriveAlarm ,ET:= m_tNotArriveCurrentTime );
(*//下料超时报警*)
m_tonUnloadAlam(IN:= iStep=4,PT:=ConveyorMotor.tUnloadAlarmDelay,Q:= ConveyorMotor.xUnloadAlarm,ET:=m_tUnloadTimer );
(*//限位报警,进料检测开关失效*)
set(  ( ((ConveyorMotor.xloadCCW AND NOT ConveyorMotor.xNegLimit)            (*反转上料，碰到负限位*)
			OR  ( NOT ConveyorMotor.xloadCCW AND NOT ConveyorMotor.xPosLimit)) (*正转上料，碰到正限位*)
		AND iStep=2) (*上料过程*)
	OR
	( iStep=4 (*下料过程*)
		AND( (ConveyorMotor.xUnloadCCW AND NOT ConveyorMotor.xPosLimit)  
			OR (NOT ConveyorMotor.xUnloadCCW AND NOT ConveyorMotor.xNegLimit)))  ,  
	ConveyorMotor.xLimitAlarrm );
mov( ( ((ConveyorMotor.xloadCCW AND NOT ConveyorMotor.xNegLimit)            (*反转上料，碰到负限位*)
			OR  ( NOT ConveyorMotor.xloadCCW AND NOT ConveyorMotor.xPosLimit)) (*正转上料，碰到正限位*)
		AND iStep=2) (*上料过程*)
	OR
	( iStep=4 (*下料过程*)
		AND( (ConveyorMotor.xUnloadCCW AND NOT ConveyorMotor.xPosLimit)  
			OR (NOT ConveyorMotor.xUnloadCCW AND NOT ConveyorMotor.xNegLimit)))  ,
	0,
	iStep);
(*//超宽报警*)
set( (iStep=3 OR iStep=1) AND (NOT ConveyorMotor.xNegLimit OR NOT ConveyorMotor.xPosLimit) , ConveyorMotor.xOverWidthAlarm  );
(*//尺寸不足报警*)
(*//有料状态下检测两个开关都要有信号*)
set( iStep=3 AND ConveyorMotor.xSizeDeficientDetect AND (NOT ConveyorMotor.xCCWPresent OR NOT ConveyorMotor.xCWPresent) ,  ConveyorMotor.xOverWidthAlarm );
mov( iStep=3 AND ConveyorMotor.xSizeDeficientDetect AND (NOT ConveyorMotor.xCCWPresent OR NOT ConveyorMotor.xCWPresent),0,iStep);
(*//总报警*)
ConveyorMotor.xError:=ConveyorMotor.xLimitAlarrm
					OR ConveyorMotor.xNotArriveAlarm
					OR ConveyorMotor.xUnloadAlarm                                             
					OR ConveyorMotor.xOverWidthAlarm;

